
   #AUX_rgtOUT_tDriveData.iLiveCounter := #AUX_rgtOUT_tDriveData.iLiveCounter + 1;
   #AUX_rgtOUT_tDriveData.rgxControlBits.xFaultReset := #AUX_tOutputDrive.rgxControlBits.xFaultReset;
   #AUX_rgtOUT_tDriveData.rgxControlBits.xEnableBridge := #AUX_tOutputDrive.rgxControlBits.xEnableBridge;
   #AUX_rgtOUT_tDriveData.rgxControlBits.xDisableBridge := #AUX_tOutputDrive.rgxControlBits.xDisableBridge;
END_REGION

REGION Network 39 (SCL): Update data to inverter
   IF #PH_xWriteModbus THEN
   #AUX_rgdParameterArray[20] := #AUX_rgtOUT_tDriveData.dBridgeAngle_degre_10000;
   #AUX_rgdParameterArray[21] := #AUX_rgtOUT_tDriveData.dHeadDownPos_dmm;
   #AUX_rgdParameterArray[22] := #AUX_rgtOUT_tDriveData.dHeadRisePos_dmm;
   #AUX_rgdParameterArray[19] := INT_TO_DINT(#AUX_rgtOUT_tDriveData.iReturnSpeed_rpm);
   #AUX_rgdParameterArray[11] := INT_TO_DINT(#AUX_rgtOUT_tDriveData.iTimeHeadDown_ms);
   #AUX_rgdParameterArray[12] := INT_TO_DINT(#AUX_rgtOUT_tDriveData.iTimeHeadUp_ms);
   #AUX_rgdParameterArray[13] := INT_TO_DINT(#AUX_rgtOUT_tDriveData.iLubAdvanceTime_ms);
   #AUX_rgdParameterArray[14] := INT_TO_DINT(#AUX_rgtOUT_tDriveData.iLubDelayTime_ms);
   #AUX_rgdParameterArray[15] := INT_TO_DINT(#AUX_rgtOUT_tDriveData.iTimeHeadAct_ms);
   #AUX_rgdParameterArray[16] := INT_TO_DINT(#AUX_rgtOUT_tDriveData.iTimeHeadDeactiv_ms);
   #AUX_rgdParameterArray[25] := #AUX_rgtOUT_tDriveData.dPressure_mN;
   #AUX_rgdParameterArray[26] := #AUX_rgtOUT_tDriveData.dMissionID;
   #AUX_rgdParameterArray[27] := #AUX_rgtOUT_tDriveData.dMissionCounter;
   #AUX_rgdParameterArray[28] := #AUX_rgtOUT_tDriveData.dSyncroCounter;
   #AUX_rgdParameterArray[17] := INT_TO_DINT(#AUX_rgtOUT_tDriveData.iLiveCounter);
   GATHER(IN:=#AUX_rgtOUT_tDriveData.rgxControlBits,
          OUT=> #TMP_dwValue);
   #AUX_rgdParameterArray[18] := DWORD_TO_DINT(#TMP_dwValue);
   #AUX_rgdParameterArray[23] := 0;
   #AUX_rgdParameterArray[24] := 0;
   END_IF;
END_REGION
END_FUNCTION_BLOCK

FUNCTION_BLOCK "FB_CrossCutsModbusExchange_V1.00"   // FB8, LAD
TITLE = Cross cut machine V1.00
{ S7_Optimized_Access := 'TRUE' }
VERSION : 0.1
   VAR_INPUT
      IN_xGeneralReset : Bool;   // General reset
      IN_dMachineIndex : DInt;   // Tracking machine index
   END_VAR
   VAR_IN_OUT
      INO_tXcut : "FB_CrossCutsModbus_V1.00";   // Xcut DB
      INO_tMBClient : MB_CLIENT;   // MB client
      INO_stConnect : TCON_IP_v4;   // Modbus connection parameters
   END_VAR
   VAR_TEMP
      TMP_iModbus_mode : UDInt;   // Modbus mode (0=read, 1=write)
      TMP_dModbus_address : UDInt;   // Modbus address
      TMP_dModbus_length : UDInt;   // Modbus data length
      TMP_dValue : DInt;   // Modbus data length
      TMP_dIndex : DInt;   // Modbus data length
   END_VAR
   VAR CONSTANT
      CONST_DREACTTIMETRACK_MS : DInt := 50;   // Tracking machine reaction time [ms]
      CONST_DMODECUT_OPERATOR : DInt := 1;   // Cut modality - By operator
      CONST_DMODECUT_GROSS : DInt := 2;   // Cut modality - Gross width
      CONST_DMODECUT_NET : DInt := 3;   // Cut modality - Net width
      CONST_DMODECUT_YCUT : DInt := 4;   // Cut modality - YCut
      CONST_DMINCUTRANGE_CMM : DInt := 25000;   // Minimum cutting start position [mm/100]
      CONST_DMAXCUTRANGE_CMM : DInt := 500000;   // Maximum cutting start position [mm/100]
      CONST_DMAXMISSIONNUM : DInt := 1000;   // Maximum number of mission to XCUT
      CONST_DMAXWAITFEEDBACK_CMM : DInt := 20000;   // Waiting space feedback [mm/100]
      CONST_DDISABLED : DInt := 1;   // Disabled
      CONST_DENABLED : DInt := 3;   // Enabled
      CONST_DSIZEALARMS : UDInt := 32;   // Number of bool on alarms structure
      CONST_DTIMEOUTINVERTER_MS : Time := T#2000ms;   // Inverter counter timeout
      CONST_DMAXRETSPEED_RPM : DInt := 3750;   // Maximum return speed [rpm]
      CONST_DSPEED_CMM_S : DInt := 500000;   // Return travel speed [mm/100/s]
      CONST_DRAMP_CMM_S2 : DInt := 1200000;   // Return travel ramp [mm/100/s]
      CONST_DBREAKDOWNOFF_CMM : DInt := 50000;   // Break downstream offset [mm/100]
      CONST_DBREAKUPOFF_CMM : DInt := 50000;   // Break upstream offset [mm/100]
      CONST_DADDRESSMENU_READ : UDInt := 2001;   // Parameter menu start (#20.01=2001)
      CONST_DADDRESSMENU_WRITE : UDInt := 2010;   // Parameter menu start (#20.01=2001)
   END_VAR
   VAR_TEMP   // added for the SCL form of the ladder/FBD networks
      _w1 : Bool;
      _w2 : Bool;
   END_VAR
BEGIN

REGION Network 1: ####_CONSTANTS_####
END_REGION

REGION Network 2: ####_MATCH_####
END_REGION

REGION Network 3: ####_PHASES_&_LOGICS_MODBUS_####
END_REGION

REGION Network 4 (SCL): Modbus address
   IF #INO_tXcut.PH_xWriteModbus OR #INO_tXcut.PH_xEndWriteModbus THEN
       #TMP_dModbus_address := 400000 + #CONST_DADDRESSMENU_WRITE + 16384;
       #TMP_dModbus_length := 40;
       #TMP_iModbus_mode := 1;
       #TMP_dValue := 9;

   ELSE
       #TMP_dModbus_address := 400000 + #CONST_DADDRESSMENU_READ + 16384;
       #TMP_dModbus_length := 80;
       #TMP_iModbus_mode := 0;
       #TMP_dValue := 0;

   END_IF;

   FOR #TMP_dIndex := 0 TO 20 DO
       "DB_ExchangeDataModbusWrite".DataXcut[#IN_dMachineIndex].Data[#TMP_dIndex] := #INO_tXcut.AUX_rgdParameterArray[#TMP_dIndex+9];
   END_FOR;
END_REGION

REGION Network 5: MB client
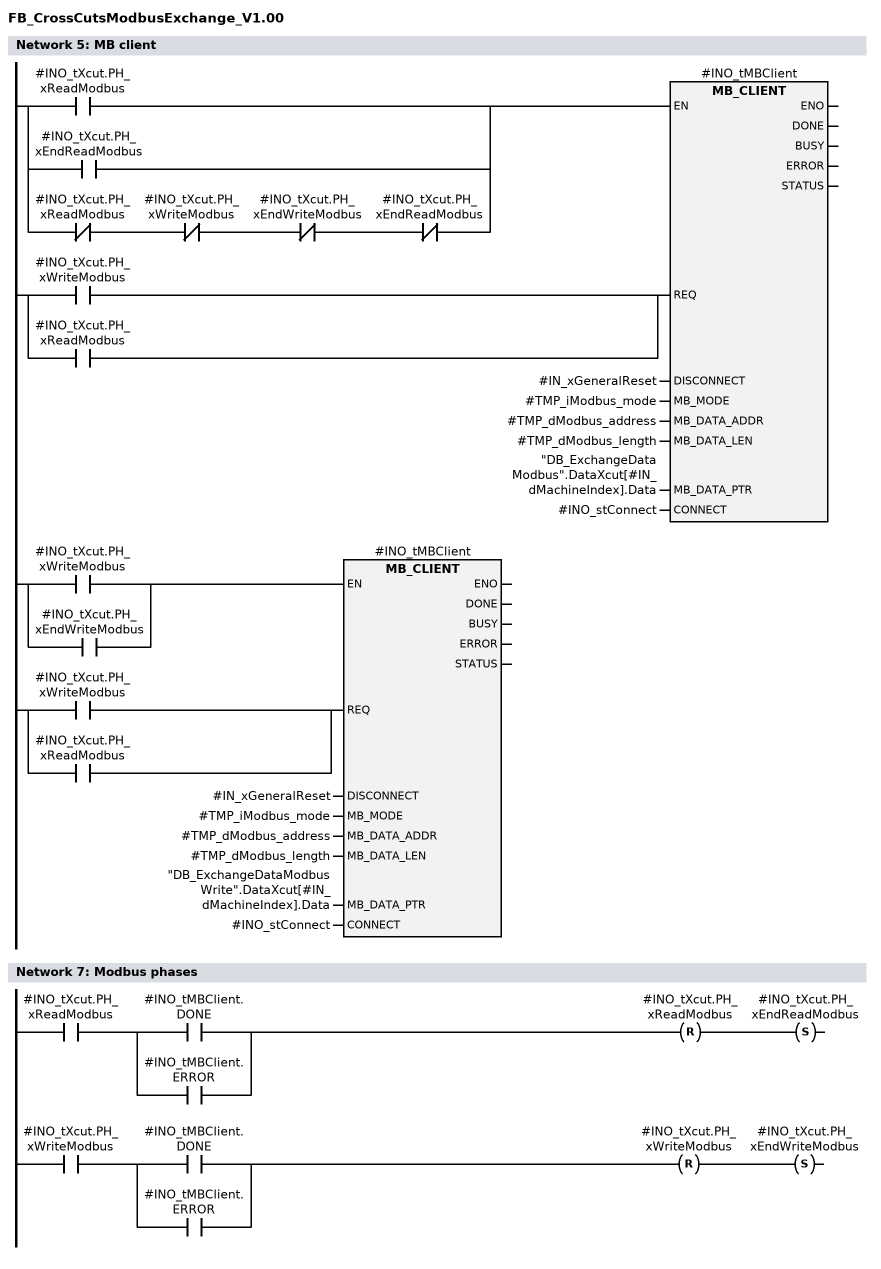
   IF #INO_tXcut.PH_xReadModbus OR #INO_tXcut.PH_xEndReadModbus OR (NOT #INO_tXcut.PH_xReadModbus AND NOT #INO_tXcut.PH_xWriteModbus AND NOT #INO_tXcut.PH_xEndWriteModbus AND NOT #INO_tXcut.PH_xEndReadModbus) THEN
       #INO_tMBClient(REQ := #INO_tXcut.PH_xWriteModbus OR #INO_tXcut.PH_xReadModbus,   // MB_CLIENT
                      DISCONNECT := #IN_xGeneralReset,
                      MB_MODE := #TMP_iModbus_mode,
                      MB_DATA_ADDR := #TMP_dModbus_address,
                      MB_DATA_LEN := #TMP_dModbus_length,
                      MB_DATA_PTR := "DB_ExchangeDataModbus".DataXcut[#IN_dMachineIndex].Data,
                      CONNECT := #INO_stConnect);
   END_IF;
   IF #INO_tXcut.PH_xWriteModbus OR #INO_tXcut.PH_xEndWriteModbus THEN
       #INO_tMBClient(REQ := #INO_tXcut.PH_xWriteModbus OR #INO_tXcut.PH_xReadModbus,   // MB_CLIENT
                      DISCONNECT := #IN_xGeneralReset,
                      MB_MODE := #TMP_iModbus_mode,
                      MB_DATA_ADDR := #TMP_dModbus_address,
                      MB_DATA_LEN := #TMP_dModbus_length,
                      MB_DATA_PTR := "DB_ExchangeDataModbusWrite".DataXcut[#IN_dMachineIndex].Data,
                      CONNECT := #INO_stConnect);
   END_IF;
END_REGION

REGION Network 6 (SCL): Array of xcut parameters (menu 20)
   IF #INO_tXcut.PH_xReadModbus AND #INO_tMBClient.DONE THEN
       #INO_tXcut.AUX_rgdParameterArray := "DB_ExchangeDataModbus".DataXcut[#IN_dMachineIndex].Data;

   END_IF;
END_REGION

REGION Network 7: Modbus phases
   RUNG wire#powerrail
      Contact( #INO_tXcut.PH_xReadModbus )
      wire#w1
      Contact( #INO_tMBClient.DONE )
      wire#w2
      R_Coil( #INO_tXcut.PH_xReadModbus )
      S_Coil( #INO_tXcut.PH_xEndReadModbus )
   END_RUNG
   RUNG wire#w1
      Contact( #INO_tMBClient.ERROR )
   END_RUNG wire#w2
   RUNG wire#powerrail
      Contact( #INO_tXcut.PH_xWriteModbus )
      wire#w3
      Contact( #INO_tMBClient.DONE )
      wire#w4
      R_Coil( #INO_tXcut.PH_xWriteModbus )
      S_Coil( #INO_tXcut.PH_xEndWriteModbus )
   END_RUNG
   RUNG wire#w3
      Contact( #INO_tMBClient.ERROR )
   END_RUNG wire#w4
   // the same network as SCL:
   #_w1 := #INO_tXcut.PH_xReadModbus AND (#INO_tMBClient.DONE OR #INO_tMBClient.ERROR);
   IF #_w1 THEN
       #INO_tXcut.PH_xReadModbus := FALSE;
       #INO_tXcut.PH_xEndReadModbus := TRUE;
   END_IF;
   #_w2 := #INO_tXcut.PH_xWriteModbus AND (#INO_tMBClient.DONE OR #INO_tMBClient.ERROR);
   IF #_w2 THEN
       #INO_tXcut.PH_xWriteModbus := FALSE;
       #INO_tXcut.PH_xEndWriteModbus := TRUE;
   END_IF;
END_REGION
END_FUNCTION_BLOCK

FUNCTION_BLOCK "FB_CrossCutOpt_V1.00"   // FB35, FBD
{ S7_Optimized_Access := 'TRUE' }
VERSION : 0.1
   VAR_INPUT
      IN_dXCutCallIndex : DInt;   // Cross cut call index
      IN_xNewTargetCall : Bool;   // New target line call request
      IN_dCapIndexCall : DInt;   // Cap Index call
      IN_xRescueCall : Bool;   // Rescue call (verify if target is still available)
      IN_dActualNumOfXCuts : DInt;   // Actual number of XCuts
      IN_rgxCutsAvailable : Array[0.."DMAXXHEADS_IND"] of Bool;   // XCut available list
      IN_rgdPiorityList : Array[0.."DMAXXHEADS_IND"] of DInt;   // Priority list value
      IN_rgdCutTime_ms : Array[0.."DMAXXHEADS_IND"] of DInt;   // Actual cutting time [ms]
   END_VAR
   VAR_IN_OUT
      INO_tOBInit : "GP_OB_Initialize";   // OB Initialize
      INO_tTrack : "UDT_CapData_Tracking";   // Tracking plate
   END_VAR
   VAR
      AUX_rgdRunningTime_ms : Array[0.."DMAXXHEADS_IND"] of DInt;   // Running time [ms]
      AUX_rgdLastExecutionTime_ms : Array[0.."DMAXXHEADS_IND"] of DInt;   // Last execution time [ms]
   END_VAR
   VAR RETAIN
      tHMR : Struct   // HMI Write data
         xEnabledPriority : Bool;   // Enabled/disable priority (1=enabled) {X|X|X|X|O}
      END_STRUCT;
      tHMW : Struct   // HMI Write data
         xEnDisPriority : Bool;   // Enable/disable priority (1=enabled) {X|X|X|X|O}
      END_STRUCT;
   END_VAR
   VAR_TEMP
      TMP_dIndex : DInt;
      TMP_dSelXCutIndex : DInt;
      TMP_dSelXCutLastUsed_ms : DInt;
      TMP_dSelXCutRunTime_ms : DInt;
      TMP_dSelXCutPrio : DInt;
   END_VAR
BEGIN

REGION Network 2 (SCL): Choose the best xcut
   IF  #IN_dXCutCallIndex = 0 AND #IN_xNewTargetCall  THEN

       #TMP_dSelXCutIndex := -1;
       #TMP_dSelXCutLastUsed_ms := 0;
       #TMP_dSelXCutRunTime_ms := 999999;
       #TMP_dSelXCutPrio := -1;
       #TMP_dIndex := 0;

       WHILE (#TMP_dIndex < #IN_dActualNumOfXCuts) DO

           //Assign xcut 1 as best
           IF #TMP_dSelXCutIndex = -1 THEN

               #TMP_dSelXCutIndex := #TMP_dIndex;
               #TMP_dSelXCutLastUsed_ms := #AUX_rgdLastExecutionTime_ms[#TMP_dIndex];
               #TMP_dSelXCutRunTime_ms := #AUX_rgdRunningTime_ms[#TMP_dIndex];
               #TMP_dSelXCutPrio := #IN_rgdPiorityList[#TMP_dIndex];

           ELSE

               IF #IN_rgxCutsAvailable[#TMP_dIndex] THEN //if xcut is enabled
                   //check if best run time is less then next cut, if not assign the cut to next
                   IF #TMP_dSelXCutRunTime_ms > #AUX_rgdRunningTime_ms[#TMP_dIndex] THEN

                       #TMP_dSelXCutIndex := #TMP_dIndex;
                       #TMP_dSelXCutLastUsed_ms := #AUX_rgdLastExecutionTime_ms[#TMP_dIndex];
                       #TMP_dSelXCutRunTime_ms := #AUX_rgdRunningTime_ms[#TMP_dIndex];
                       #TMP_dSelXCutPrio := #IN_rgdPiorityList[#TMP_dIndex];


                   ELSIF #TMP_dSelXCutRunTime_ms = #AUX_rgdRunningTime_ms[#TMP_dIndex] THEN
                       //if run time is the same assign the cut to highest priority bridge
                       IF #TMP_dSelXCutPrio < #IN_rgdPiorityList[#TMP_dIndex] THEN
                           #TMP_dSelXCutIndex := #TMP_dIndex;
                           #TMP_dSelXCutLastUsed_ms := #AUX_rgdLastExecutionTime_ms[#TMP_dIndex];
                           #TMP_dSelXCutRunTime_ms := #AUX_rgdRunningTime_ms[#TMP_dIndex];
                           #TMP_dSelXCutPrio := #IN_rgdPiorityList[#TMP_dIndex];

                        //if priority is the same assign cut to the one which has been waiting for a longer time   
                       ELSIF #TMP_dSelXCutPrio = #IN_rgdPiorityList[#TMP_dIndex] THEN

                           IF #TMP_dSelXCutLastUsed_ms < #AUX_rgdLastExecutionTime_ms[#TMP_dIndex] THEN
                               #TMP_dSelXCutIndex := #TMP_dIndex;
                               #TMP_dSelXCutLastUsed_ms := #AUX_rgdLastExecutionTime_ms[#TMP_dIndex];
                               #TMP_dSelXCutRunTime_ms := #AUX_rgdRunningTime_ms[#TMP_dIndex];
                               #TMP_dSelXCutPrio := #IN_rgdPiorityList[#TMP_dIndex];

                           END_IF;
                       END_IF;
                   END_IF;

               END_IF;
           END_IF;
           #TMP_dIndex += 1;
       END_WHILE;

       //Associate the relative XCut
       IF #TMP_dSelXCutIndex > -1 THEN

           #AUX_rgdRunningTime_ms[#TMP_dSelXCutIndex] := #IN_rgdCutTime_ms[#TMP_dSelXCutIndex ];
           #AUX_rgdLastExecutionTime_ms[#TMP_dSelXCutIndex] := 0;
           #INO_tTrack.rgtTrackCaps[#IN_dCapIndexCall].tCap.tRequests.rgbXCutPrioSelect[#TMP_dSelXCutIndex] := 1;
       END_IF;


   END_IF;
END_REGION

REGION Network 3 (SCL): Decrement counters only the first call
   IF #IN_dXCutCallIndex = 0 THEN

       FOR #TMP_dIndex := 0 TO "DMAXXHEADS_IND" DO

           #AUX_rgdRunningTime_ms[#TMP_dIndex] -= #INO_tOBInit.OUT_dExecutionTime_ms;
           #AUX_rgdLastExecutionTime_ms[#TMP_dIndex] += #INO_tOBInit.OUT_dExecutionTime_ms;

           IF #AUX_rgdRunningTime_ms[#TMP_dIndex] < 0 THEN
               #AUX_rgdRunningTime_ms[#TMP_dIndex] := 0;                        
           END_IF;            

           IF #AUX_rgdLastExecutionTime_ms[#TMP_dIndex] > 3600000 THEN
               #AUX_rgdLastExecutionTime_ms[#TMP_dIndex] := 3600000;
           END_IF;

       END_FOR;

   END_IF;
END_REGION
END_FUNCTION_BLOCK

// folder: 03_Programs_Logics/MCC1200/04_Encoder

FUNCTION_BLOCK "FB_Digitizer_V1.00"   // FB3, LAD
{ S7_Optimized_Access := 'TRUE' }
VERSION : 0.1
   VAR_INPUT
      IN_xCycleON : Bool;   // Cycle ON
      IN_xCycleONDel : Bool;   // Delayed cycle ON signal
      IN_xGeneralReset : Bool;   // General reset
      IN_xResetAlarms : Bool;   // Reset alarms
      IN_xFaultsEnabled : Bool;   // Faults enabled
      IN_tInterfaceID : Hw_Any;   // Interface ID
      IN_tID : Conn_Ouc;   // Connection ID
      IN_tRemoteAddress : IP_V4;   // Remote IP address
      IN_uiRemotePort : UInt;   // Remote port
      INPUTS : Struct
         xGlassPresence : Bool;   // INPUT.Photocell glass presence
         dEncCounter_count : DInt;   // INPUT.Encoder counter [count]
      END_STRUCT;
      IN_xSimulationActive : Bool;   // Enable simulation (EXPERT USER)
   END_VAR
   VAR_OUTPUT
      OUTPUTS : Struct   // Outputs
         xDescentEncoder : Bool;   // OUTPUT.Descent encoder
         xCounterSWGate : Bool;   // OUTPUT.Card software gate
      END_STRUCT;
   END_VAR
   VAR_IN_OUT
      INO_tEnc : "UDT_Encoder";   // Encoder data
   END_VAR
   VAR RETAIN
      tHMR : Struct
         xMan_DescEncFdbk : Bool;   // Manual mode. Feedback descent encoder
         dEncoderStatus : DInt;   // Encoder status (1=Stop 3=Running 7=Anomaly)
         dCalibrationF1Unit_unit : DInt;   // Calibration actual F1 [unit]
         dCalibrationF2Unit_unit : DInt;   // Calibration actual F2 [unit]
         dActualEncoderSpeed_mm_min : DInt;   // Actual encoder speed [mm/min]
         dFm152Status : DInt;   // Status of the Fm152 card
         dCalibrationCardF1Unit_unit : DInt;   // Calibration actual F1 read from FM [unit]
         xManComEn : Bool;   // Manual command enabled
         dCalibrationCardF2Unit_unit : DInt;   // Calibration actual F2 read from FM [unit]
      END_STRUCT;
      tHMW : Struct
         xCalibUpdateF1 : Bool;   // Calibration update F1 value
         xCalibUpdateF2 : Bool;   // Calibration update F2 value
         xCalibRequest : Bool;   // Calibration length request
         xMan_DescentEnc : Bool;   // Manual encoder descent
         xGlassSensorEnabled : Bool;   // Glass presence sensor are enabled
         dCalibTheoLength_cmm : DInt;   // Calibration theorical length [mm/100]
         dCalibRealLength_cmm : DInt;   // Calibration real length [mm/100]
         dCalibWriteF1_unit : DInt;   // Calibration write F1 [unit]
         dCalibWriteF2_unit : DInt;   // Calibration write F2 [unit]
         dRequestJogSpeed_mm_min : DInt;   // Jog speed requested [mm/min]
         xEnDisManCom : Bool;   // Enable disable manual command
      END_STRUCT;
   END_VAR
   VAR
      tALM : Struct   // HMI Alarms
         tS : Struct   // Stopping faults
            xNoEncPulses : Bool;   // BQ.No encoder pulses
            xSpeedOutLimits : Bool;   // BQ.Speed outside min max limits
            xSpare_2 : Bool;
            xSpare_3 : Bool;
            xSpare_4 : Bool;
            xSpare_5 : Bool;
            xSpare_6 : Bool;
            xSpare_7 : Bool;
            xSpare_8 : Bool;
            xSpare_9 : Bool;
            xSpare_10 : Bool;
            xSpare_11 : Bool;
            xSpare_12 : Bool;
            xSpare_13 : Bool;
            xSpare_14 : Bool;
            xSpare_15 : Bool;
            xSpare_16 : Bool;
            xSpare_17 : Bool;
            xSpare_18 : Bool;
            xSpare_19 : Bool;
            xSpare_20 : Bool;
            xSpare_21 : Bool;
            xSpare_22 : Bool;
            xSpare_23 : Bool;
            xSpare_24 : Bool;
            xSpare_25 : Bool;
            xSpare_26 : Bool;
            xSpare_27 : Bool;
            xSpare_28 : Bool;
            xSpare_29 : Bool;
            xSpare_30 : Bool;
            xSpare_31 : Bool;
         END_STRUCT;
         tF : Struct   // Faults
            xMissingEncPulses : Bool;   // Missing encoder pulses
            xFm152SendError : Bool;   // FM152. Sending data error
            xFm152SendTimeout : Bool;   // FM152. Sending data timeout
            xFm152RecvTimeout : Bool;   // FM152.Receiving data timeout
            xSpare_4 : Bool;
            xSpare_5 : Bool;
            xSpare_6 : Bool;
            xSpare_7 : Bool;
            xSpare_8 : Bool;
            xSpare_9 : Bool;
            xSpare_10 : Bool;
            xSpare_11 : Bool;
            xSpare_12 : Bool;
            xSpare_13 : Bool;
            xSpare_14 : Bool;
            xSpare_15 : Bool;
            xSpare_16 : Bool;
            xSpare_17 : Bool;
            xSpare_18 : Bool;
            xSpare_19 : Bool;
            xSpare_20 : Bool;
            xSpare_21 : Bool;
            xSpare_22 : Bool;
            xSpare_23 : Bool;
            xSpare_24 : Bool;
            xSpare_25 : Bool;
            xSpare_26 : Bool;
            xSpare_27 : Bool;
            xSpare_28 : Bool;
            xSpare_29 : Bool;
            xSpare_30 : Bool;
            xSpare_31 : Bool;
         END_STRUCT;
         tW : Struct   // Warnings
            xSpare_0 : Bool;
            xSpare_1 : Bool;
            xSpare_2 : Bool;
            xSpare_3 : Bool;
            xSpare_4 : Bool;
            xSpare_5 : Bool;
            xSpare_6 : Bool;
            xSpare_7 : Bool;
            xSpare_8 : Bool;
            xSpare_9 : Bool;
            xSpare_10 : Bool;
            xSpare_11 : Bool;
            xSpare_12 : Bool;
            xSpare_13 : Bool;
            xSpare_14 : Bool;
            xSpare_15 : Bool;
            xSpare_16 : Bool;
            xSpare_17 : Bool;
            xSpare_18 : Bool;
            xSpare_19 : Bool;
            xSpare_20 : Bool;
            xSpare_21 : Bool;
            xSpare_22 : Bool;
            xSpare_23 : Bool;
            xSpare_24 : Bool;
            xSpare_25 : Bool;
            xSpare_26 : Bool;
            xSpare_27 : Bool;
            xSpare_28 : Bool;
            xSpare_29 : Bool;
            xSpare_30 : Bool;
            xSpare_31 : Bool;
         END_STRUCT;
      END_STRUCT;
      AUX_dTimePhotoWheel_ms : DInt;   // Time from photocell and encoder wheel [ms]
      ST_xEncDownPosition : Bool;   // Encoder is in down position
      ST_xStoppingFaults : Bool;   // Stopping faults
      ST_xFaults : Bool;   // Faults
      ST_xOuputEnable : Bool;   // Output enable
      OUT_xDescentEncoder : Bool;   // Output copy descent encoder
      tmON_DescentEnc : TON_TIME;   // Timer TON for waiting descent encoder
      tmON_EncReactTime : TON_TIME;   // Timer TON encoder reaction time
      tmON_GlassOnEncDel : TON_TIME;   // Timer TON glass under encoder
      tmON_TimeoutSendData : TON_TIME;   // Timer TON sending data
      ST_xGlassUnderEnc : Bool;   // Glass present under the encoder
      ST_xEncDescReq : Bool;   // Encoder descent request
      AUX_lrTimingCounter_s : LReal;   // Timing counter [s]
      AUX_lrElapsedTime_s : LReal;   // Elapsed time from previous call [s]
      AUX_lrRuntimeMemory_s : LReal;   // Variable used for runtime instruction [s]
      AUX_dLastCounterValueFast_cmm : DInt;   // Last counter value fast [mm/100]
      AUX_dLastCounterValue_cmm : DInt;   // Last counter value [mm/100]
      FB_TSend : TSEND_C;
      AUX_tFM152SndReadSt : Struct   // FM152 read status request
         bEOT : Byte;   // Eot
         bAD1 : Byte;   // Ad1
         bAD2 : Byte;   // Ad2
         bC1 : Byte;   // C1
         bC2 : Byte;   // C2
         bENQ : Byte;   // Enq
      END_STRUCT;
      AUX_tFM152SndReadF1 : Struct   // FM152 read F1 request
         bEOT : Byte;   // Eot
         bAD1 : Byte;   // Ad1
         bAD2 : Byte;   // Ad2
         bC1 : Byte;   // C1
         bC2 : Byte;   // C2
         bENQ : Byte;   // Enq
      END_STRUCT;
      AUX_tFM152SndReadF2 : Struct   // FM152 read F2 request
         bEOT : Byte;   // Eot
         bAD1 : Byte;   // Ad1
         bAD2 : Byte;   // Ad2
         bC1 : Byte;   // C1
         bC2 : Byte;   // C2
         bENQ : Byte;   // Enq
      END_STRUCT;
      AUX_tFM152SndWriteF1 : Struct   // FM152 write F1 request
         bEOT : Byte;   // Eot
         bAD1 : Byte;   // Ad1
         bAD2 : Byte;   // Ad2
         bSTX : Byte;   // Stx
         bC1 : Byte;   // C1
         bC2 : Byte;   // C2
         bVal1 : Byte;   // Value char 1
         bVal2 : Byte;   // Value char 2
         bVal3 : Byte;   // Value char 3
         bVal4 : Byte;   // Value char 4
         bVal5 : Byte;   // Value char 5
         bETX : Byte;   // Etx
         bBCC : Byte;   // Bcc
      END_STRUCT;
      AUX_tFM152SndWriteF2 : Struct   // FM152 write F2 request
         bEOT : Byte;   // Eot
         bAD1 : Byte;   // Ad1
         bAD2 : Byte;   // Ad2
         bSTX : Byte;   // Stx
         bC1 : Byte;   // C1
         bC2 : Byte;   // C2
         bVal1 : Byte;   // Value char 1
         bVal2 : Byte;   // Value char 2
         bVal3 : Byte;   // Value char 3
         bVal4 : Byte;   // Value char 4
         bVal5 : Byte;   // Value char 5
         bETX : Byte;   // Etx
         bBCC : Byte;   // Bcc
      END_STRUCT;
      AUX_tFM152SndWriteJog : Struct   // FM152 write jog request
         bEOT : Byte;   // Eot
         bAD1 : Byte;   // Ad1
         bAD2 : Byte;   // Ad2
         bSTX : Byte;   // Stx
         bC1 : Byte;   // C1
         bC2 : Byte;   // C2
         bVal1 : Byte;   // Value char 1
         bVal2 : Byte;   // Value char 2
         bVal3 : Byte;   // Value char 3
         bVal4 : Byte;   // Value char 4
         bVal5 : Byte;   // Value char 5
         bETX : Byte;   // Etx
         bBCC : Byte;   // Bcc
      END_STRUCT;
      AUX_tFM152SndWriteRampRef : Struct   // FM152 write ramp reference
         bEOT : Byte;   // Eot
         bAD1 : Byte;   // Ad1
         bAD2 : Byte;   // Ad2
         bSTX : Byte;   // Stx
         bC1 : Byte;   // C1
         bC2 : Byte;   // C2
         bC3 : Byte;   // C3
         bC4 : Byte;   // C4
         bETX : Byte;   // Etx
         bBCC : Byte;   // Bcc
      END_STRUCT;
      AUX_tFM152SndWriteRampJog : Struct   // FM152 write ramp jog reference
         bEOT : Byte;   // Eot
         bAD1 : Byte;   // Ad1
         bAD2 : Byte;   // Ad2
         bSTX : Byte;   // Stx
         bC1 : Byte;   // C1
         bC2 : Byte;   // C2
         bC3 : Byte;   // C3
         bC4 : Byte;   // C4
         bETX : Byte;   // Etx
         bBCC : Byte;   // Bcc
      END_STRUCT;
      AUX_tFM152SndWriteRamp : Struct   // FM152 write ramp
         bEOT : Byte;   // Eot
         bAD1 : Byte;   // Ad1
         bAD2 : Byte;   // Ad2
         bSTX : Byte;   // Stx
         bC1 : Byte;   // C1
         bC2 : Byte;   // C2
         bC3 : Byte;   // C3
         bC4 : Byte;   // C4
         bETX : Byte;   // Etx
         bBCC : Byte;   // Bcc
      END_STRUCT;
      AUX_tFM152SndActivateData : Struct   // FM152 activate data
         bEOT : Byte;   // Eot
         bAD1 : Byte;   // Ad1
         bAD2 : Byte;   // Ad2
         bSTX : Byte;   // Stx
         bC1 : Byte;   // C1
         bC2 : Byte;   // C2
         bC3 : Byte;   // C3
         bETX : Byte;   // Etx
         bBCC : Byte;   // Bcc
      END_STRUCT;
      AUX_tFM152RecvStatus : Struct   // FM152 read status feedback
         bSTX : Byte;   // STX
         bC1 : Byte;   // C1
         bC2 : Byte;   // C2
         bC3 : Byte;   // C3
         bC4 : Byte;   // C4
         bC5 : Byte;   // C5
         bD1 : Byte;   // D1
         bD2 : Byte;   // D2
         bETX : Byte;   // ETX
         bBCC : Byte;   // BCC
      END_STRUCT;
      AUX_tFM152RecvF1 : Struct   // FM152 read F1 feedback
         bSTX : Byte;   // STX
         bC1 : Byte;   // C1
         bC2 : Byte;   // C2
         bD1 : Byte;   // D1
         bD2 : Byte;   // D2
         bD3 : Byte;   // D3
         bD4 : Byte;   // D4
         bD5 : Byte;   // D5
         bETX : Byte;   // ETX
         bBCC : Byte;   // BCC
      END_STRUCT;
      AUX_tFM152RecvF2 : Struct   // FM152 read F2 feedback
         bSTX : Byte;   // STX
         bC1 : Byte;   // C1
         bC2 : Byte;   // C2
         bD1 : Byte;   // D1
         bD2 : Byte;   // D2
         bD3 : Byte;   // D3
         bD4 : Byte;   // D4
         bD5 : Byte;   // D5
         bETX : Byte;   // ETX
         bBCC : Byte;   // BCC
      END_STRUCT;
      AUX_tFM152RecvAck : Struct   // FM152 read ACK feedback
         bACK : Byte;   // ACK
      END_STRUCT;
      AUX_dPrepTelType : DInt;   // FM152 - Prepare type of packet
      ST_xFm152PhaseProgr : Bool;   // FM152 - Phase in progress
      AUX_tConnData : TCON_IP_v4;   // FM152 - Connection data structure
      AUX_xResetSendConnection : Bool;   // FM152 - Reset the estabilished send connection
      ST_xWarnings : Bool;   // Warnings
      tPhases : Struct   // Phases
         xPrepareTelegram : Bool;   // FM152 - Prepare telegram
         xEndPrepareTelegram : Bool;   // FM152 - End prepare telegram
         xWaitingFm152Reply : Bool;   // FM152 - Waiting reply
         xEndWaitingFm152Reply : Bool;   // FM152 - End waiting reply
         xSpare4 : Bool;
         xSpare5 : Bool;
         xSpare6 : Bool;
         xSpare7 : Bool;
         xSpare8 : Bool;
         xSpare9 : Bool;
         xSpare10 : Bool;
         xSpare11 : Bool;
         xSpare12 : Bool;
         xSpare13 : Bool;
         xSpare14 : Bool;
         xSpare15 : Bool;
         xSpare16 : Bool;
         xSpare17 : Bool;
         xSpare18 : Bool;
         xSpare19 : Bool;
         xSpare20 : Bool;
         xSpare21 : Bool;
         xSpare22 : Bool;
         xSpare23 : Bool;
         xSpare24 : Bool;
         xSpare25 : Bool;
         xSpare26 : Bool;
         xSpare27 : Bool;
         xSpare28 : Bool;
         xSpare29 : Bool;
         xSpare30 : Bool;
         xSpare31 : Bool;
      END_STRUCT;
      FB_TReceive : TRCV_C;
      AUX_xResetRecvConnection : Bool;   // FM152 - Reset the estabilished receive connection
      AUX_rgbTempRecvBuffer : Array[0..19] of Byte;   // FM152 - Temporary receive buffer
      AUX_rgbReceiveBuffer : Array[0..99] of Byte;   // FM152 - Receive buffer
      AUX_dActualElBuffer : DInt;   // FM152 - Actual number of element on receive buffer
      tmON_TimeoutRecvData : TON_TIME;   // FM152 - Timeout receive data
      AUX_rgbTempSendBuffer : Array[0..19] of Byte;   // FM152 - Temporary send buffer
      AUX_dNumByteToSend : DInt;   // FM152 - Number of byte to send
      ST_xRefreshFM152 : Bool;   // FM152 - Request refresh data
      ST_xCondOkMan : Bool;   // Condition ok manual command
      AUX_dLastManualSpeed_mm_min : DInt;   // FM152 - Last manual speed [mm/min]
   END_VAR
   VAR_TEMP
      TMP_xPrepareTelegram : Bool;
      TMP_strValue : String[6];
      TMP_dwValue : DWord;
      TMP_dBufferPos : DInt;
      TMP_iRetVal : Int;
      TMP_bBBC : Byte;
      TMP_strStatus : String[2];
      TMP_xFm152ValidReply : Bool;
      TMP_strF1F2Value : String[5];
      TMP_dElapsedPulses_cmm : DInt;
      TMP_rF1Unit : Real;
      TMP_dDifferenceSpeed_mm_min : DInt;
   END_VAR
   VAR CONSTANT
      CONST_DDISTANCEPH_CMM : DInt := 30000;   // Distance of the photocell from the wheel [mm/100]
      CONST_DMAXTIMEPHOTOWHEEL_MS : DInt := 20000;   // Maximum time distance photocell to wheel [ms]
      CONST_UDSIZEALARMS : UDInt := 32;   // Number of bool on alarms structure
      CONST_DENCREACTTIME_MS : DInt := 250;   // Encoder reaction time [ms]
      CONST_DMANUAL : DInt := 1;   // Manual mode
      CONST_DAUTO : DInt := 4;   // Automatic mode
      CONST_DMANREQ : DInt := 8;   // Manual request
      CONST_DREFRESHSPEED_S : DInt := 5;   // Refresh speed time [s]
      CONST_DFM152_TEL_IDLE : DInt := 0;   // FM152 - Prepare packet idle
      CONST_DFM152_TEL_READST : DInt := 1;   // FM152 - Prepare packet read status
      CONST_DFM152_TEL_READST_NUMBYTE : DInt := 6;   // FM152 - Prepare packet read status number of byte to send
      CONST_DFM152_TEL_READF1 : DInt := 2;   // FM152 - Prepare packet read F1
      CONST_DFM152_TEL_READF1_NUMBYTE : DInt := 6;   // FM152 - Prepare packet read F1 number of byte to send
      CONST_DFM152_TEL_READF2 : DInt := 3;   // FM152 - Prepare packet read F2
      CONST_DFM152_TEL_READF2_NUMBYTE : DInt := 6;   // FM152 - Prepare packet read F2 number of byte to send
      CONST_DFM152_TEL_WRITEF1 : DInt := 4;   // FM152 - Prepare packet write F1
      CONST_DFM152_TEL_WRITEF1_NUMBYTE : DInt := 13;   // FM152 - Prepare packet write F1 number of byte to send
      CONST_DFM152_TEL_WRITEF2 : DInt := 5;   // FM152 - Prepare packet write F2
      CONST_DFM152_TEL_WRITEF2_NUMBYTE : DInt := 13;   // FM152 - Prepare packet write F2 number of byte to send
      CONST_DFM152_TEL_WRITEJOG : DInt := 6;   // FM152 - Prepare packet write jog
      CONST_DFM152_TEL_WRITEJOG_NUMBYTE : DInt := 13;   // FM152 - Prepare packet write jog number of byte to send
      CONST_DFM152_TEL_WRITERAMPREF : DInt := 7;   // FM152 - Prepare ramp reference
      CONST_DFM152_TEL_WRITERAMPREF_NUMBYTE : DInt := 10;   // FM152 - Prepare ramp reference number of byte to send
      CONST_DFM152_TEL_WRITERAMPJOG : DInt := 8;   // FM152 - Prepare ramp jog
      CONST_DFM152_TEL_WRITERAMPJOG_NUMBYTE : DInt := 10;   // FM152 - Prepare ramp jog number of byte to send
      CONST_DFM152_TEL_WRITERAMP : DInt := 9;   // FM152 - Prepare ramp
      CONST_DFM152_TEL_WRITERAMP_NUMBYTE : DInt := 10;   // FM152 - Prepare ramp number of byte to send
      CONST_DFM152_TEL_REQACTDATA : DInt := 10;   // FM152 - Request activate data
      CONST_DFM152_TEL_REQACTDATA_NUMBYTE : DInt := 9;   // FM152 - Request activate data number of byte to send
      CONST_BFM152_EOT : Byte := 16#4;   // FM152 - EOT
      CONST_BFM152_AD1 : Byte := 16#31;   // FM152 - AD1
      CONST_BFM152_AD2 : Byte := 16#31;   // FM152 - AD2
      CONST_BFM152_STX : Byte := 16#2;   // FM152 - STX
      CONST_BFM152_ETX : Byte := 16#3;   // FM152 - ETX
      CONST_BFM152_ACK : Byte := 16#6;   // FM152 - ACK
      CONST_BFM152_NACK : Byte := 16#21;   // FM152 - NACK
      CONST_BFM152_ENQ : Byte := 16#5;   // FM152 - ENQ
      CONST_BCONNTYPE : Byte := 16#0B;   // FM152 - Connection type
      CONST_DTIMEOUTSENDDATA_MS : DInt := 5000;   // FM152 - Timeout sending data [ms]
      CONST_DTIMEOUTRECVDATA_MS : DInt := 5000;   // FM152 - Timeout receive data [ms]
      CONST_DFM152_RECVSTATUSSIZE : DInt := 10;   // FM152 - Number of byte on the receive status packet
      CONST_DFM152_RECVF1F2SIZE : DInt := 10;   // FM152 - Number of byte on the receive F1 / F2 packet
      CONST_DFM152_ACK_NACKSIZE : DInt := 1;   // FM152 - Number of byre received on ACK / NACK
   END_VAR
   VAR_TEMP   // added for the SCL form of the ladder/FBD networks
      _w1 : Bool;
   END_VAR
BEGIN

REGION Network 1: ####_COSTANTS_####
END_REGION

REGION Network 2 (SCL): ### SIMULATION ###
   IF "SIMULATION_ACTIVE" THEN

       #INPUTS.dEncCounter_count := #INO_tEnc.dActualEncoderCounter_cmm;

   END_IF;
END_REGION

REGION Network 3: ####_MATCH_####
END_REGION

REGION Network 4 (SCL): FM152 - Request refresh data
   #TMP_dDifferenceSpeed_mm_min := ABS(#tHMW.dRequestJogSpeed_mm_min - #AUX_dLastManualSpeed_mm_min);

   IF (#TMP_dDifferenceSpeed_mm_min > 100) OR (#tHMR.dCalibrationCardF1Unit_unit <> #tHMR.dCalibrationF1Unit_unit)  THEN
       #ST_xRefreshFM152 := TRUE;
       #AUX_dLastManualSpeed_mm_min := #tHMW.dRequestJogSpeed_mm_min;    
   END_IF;
END_REGION

REGION Network 5: Calculate runtime execution
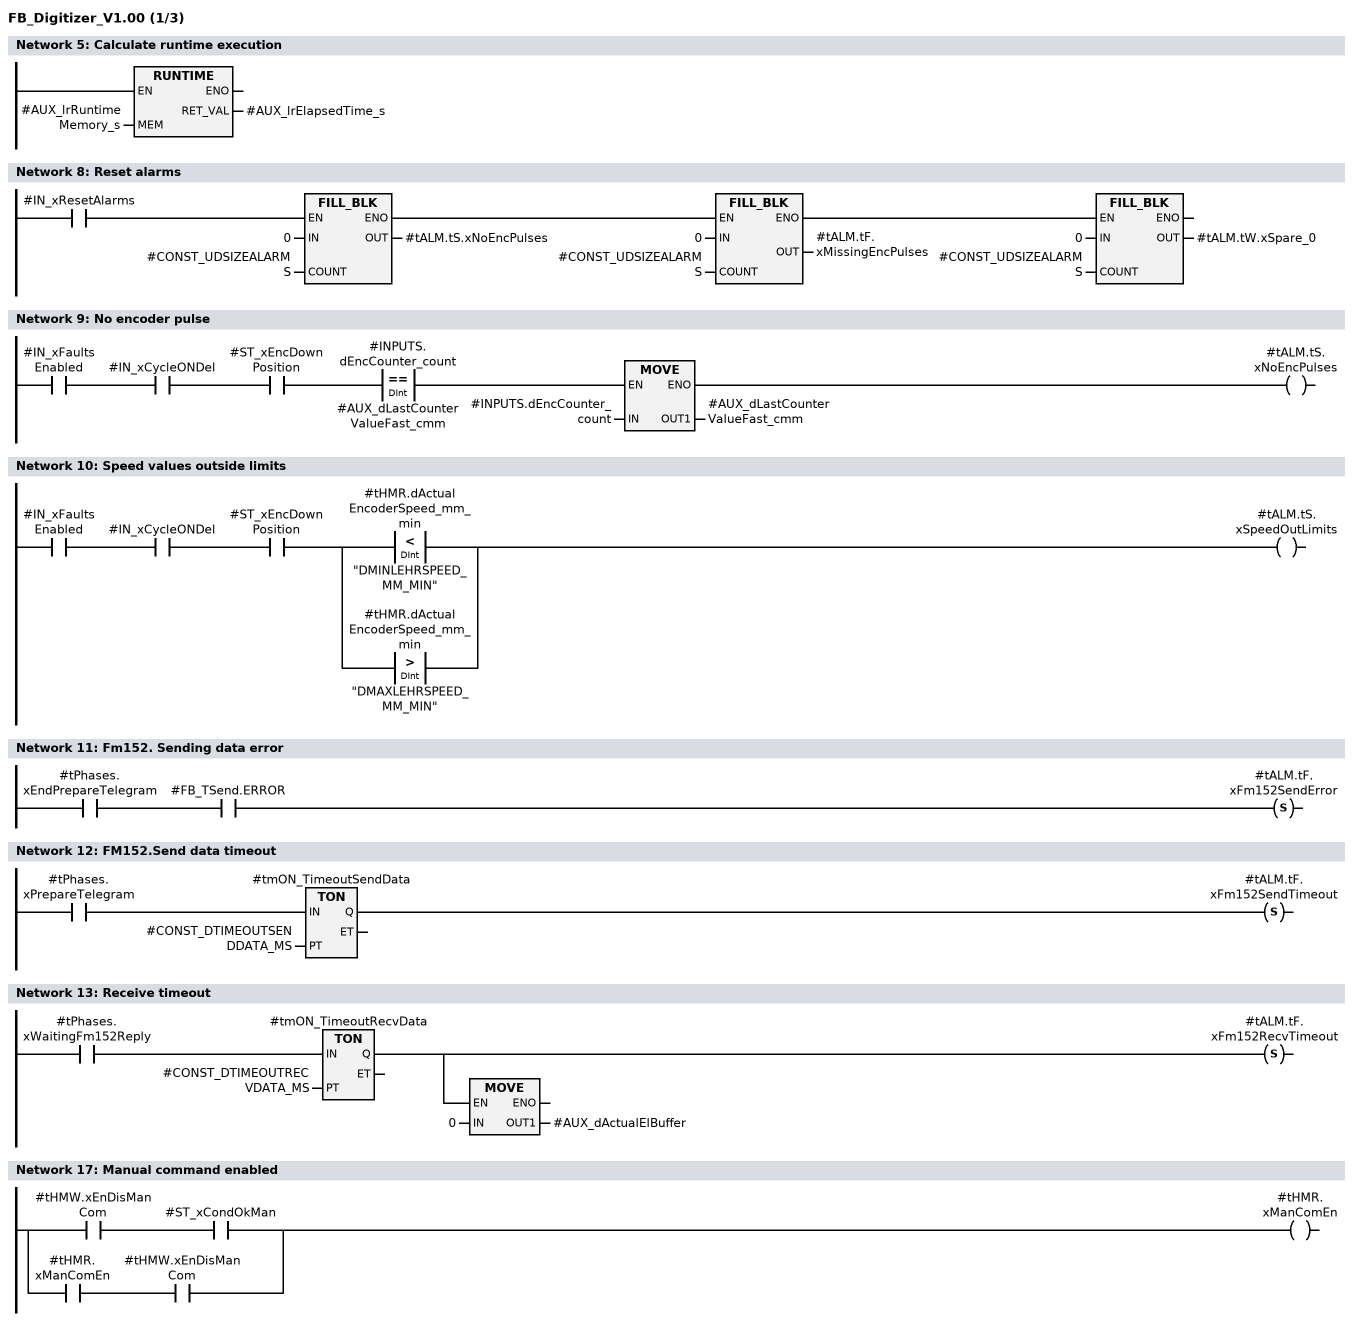
   // no SCL statement known for Runtime: written as a call
   #AUX_lrElapsedTime_s := Runtime(mem := #AUX_lrRuntimeMemory_s);
END_REGION

REGION Network 6 (SCL): Calculate time from photo to wheel
   #AUX_dTimePhotoWheel_ms := REAL_TO_DINT(DINT_TO_REAL( #CONST_DDISTANCEPH_CMM) / #INO_tEnc.rActSpeedValue_cmm_ms);

   IF #AUX_dTimePhotoWheel_ms < 0 THEN
       #AUX_dTimePhotoWheel_ms := 0;
   ELSIF #AUX_dTimePhotoWheel_ms > #CONST_DMAXTIMEPHOTOWHEEL_MS THEN
       #AUX_dTimePhotoWheel_ms := #CONST_DMAXTIMEPHOTOWHEEL_MS;
   END_IF;
END_REGION

REGION Network 7: ####_ALARMS_####
END_REGION

REGION Network 8: Reset alarms
   RUNG wire#powerrail
      Contact( #IN_xResetAlarms )
      FillBlockI(in := 0, count := #CONST_UDSIZEALARMS, out => #tALM.tS.xNoEncPulses)
      FillBlockI(in := 0, count := #CONST_UDSIZEALARMS, out => #tALM.tF.xMissingEncPulses)
      FillBlockI(in := 0, count := #CONST_UDSIZEALARMS, out => #tALM.tW.xSpare_0)
   END_RUNG
   // the same network as SCL:
   IF #IN_xResetAlarms THEN
       FILL_BLK(IN := 0, COUNT := #CONST_UDSIZEALARMS, OUT => #tALM.tS.xNoEncPulses);
       FILL_BLK(IN := 0, COUNT := #CONST_UDSIZEALARMS, OUT => #tALM.tF.xMissingEncPulses);
       FILL_BLK(IN := 0, COUNT := #CONST_UDSIZEALARMS, OUT => #tALM.tW.xSpare_0);
   END_IF;
END_REGION

